(* Logix 5000 project; controller UOWHF Emulate 5570 rev 30.12; software revision 30.00; part 6 of 13 *)
(* tags used below, declared in another part *)
   UOWHF_Add_c : DINT;
   UOWHF_Msg : DINT[16];
   UOWHF_OutputMaxInd : DINT;
   UOWHF_Result : DINT[16];
(* MainProgram, continued *)

   		UOWHF_Result[5].31:=0;
   		UOWHF_Result[6]:=UOWHF_Result[6] + 895405157+UOWHF_Add_c;
   		UOWHF_Add_c.6:=UOWHF_Result[6].31;
   		UOWHF_Result[6].31:=0;
   	End_If;
   	If UOWHF_Msg[9].[21] Then
   		UOWHF_Result[0]:=UOWHF_Result[0] + 660161237+UOWHF_Add_c;
   		UOWHF_Add_c.0:=UOWHF_Result[0].31;
   		UOWHF_Result[0].31:=0;
   		UOWHF_Result[1]:=UOWHF_Result[1] + 1315089035+UOWHF_Add_c;
   		UOWHF_Add_c.1:=UOWHF_Result[1].31;
   		UOWHF_Result[1].31:=0;
   		UOWHF_Result[2]:=UOWHF_Result[2] + 1287512548+UOWHF_Add_c;
   		UOWHF_Add_c.2:=UOWHF_Result[2].31;
   		UOWHF_Result[2].31:=0;
   		UOWHF_Result[3]:=UOWHF_Result[3] + 1179731775+UOWHF_Add_c;
   		UOWHF_Add_c.3:=UOWHF_Result[3].31;
   		UOWHF_Result[3].31:=0;
   		UOWHF_Result[4]:=UOWHF_Result[4] + 1598255528+UOWHF_Add_c;
   		UOWHF_Add_c.4:=UOWHF_Result[4].31;
   		UOWHF_Result[4].31:=0;
   		UOWHF_Result[5]:=UOWHF_Result[5] + 1383999784+UOWHF_Add_c;
   		UOWHF_Add_c.5:=UOWHF_Result[5].31;
   		UOWHF_Result[5].31:=0;
   		UOWHF_Result[6]:=UOWHF_Result[6] + 83372341+UOWHF_Add_c;
   		UOWHF_Add_c.6:=UOWHF_Result[6].31;
   		UOWHF_Result[6].31:=0;
   	End_If;
   	If UOWHF_Msg[9].[22] Then
   		UOWHF_Result[0]:=UOWHF_Result[0] + 1715876547+UOWHF_Add_c;
   		UOWHF_Add_c.0:=UOWHF_Result[0].31;
   		UOWHF_Result[0].31:=0;
   		UOWHF_Result[1]:=UOWHF_Result[1] + 985647794+UOWHF_Add_c;
   		UOWHF_Add_c.1:=UOWHF_Result[1].31;
   		UOWHF_Result[1].31:=0;
   		UOWHF_Result[2]:=UOWHF_Result[2] + 1915071159+UOWHF_Add_c;
   		UOWHF_Add_c.2:=UOWHF_Result[2].31;
   		UOWHF_Result[2].31:=0;
   		UOWHF_Result[3]:=UOWHF_Result[3] + 1355115977+UOWHF_Add_c;
   		UOWHF_Add_c.3:=UOWHF_Result[3].31;
   		UOWHF_Result[3].31:=0;
   		UOWHF_Result[4]:=UOWHF_Result[4] + 296913181+UOWHF_Add_c;
   		UOWHF_Add_c.4:=UOWHF_Result[4].31;
   		UOWHF_Result[4].31:=0;
   		UOWHF_Result[5]:=UOWHF_Result[5] + 1237257487+UOWHF_Add_c;
   		UOWHF_Add_c.5:=UOWHF_Result[5].31;
   		UOWHF_Result[5].31:=0;
   		UOWHF_Result[6]:=UOWHF_Result[6] + 1778504117+UOWHF_Add_c;
   		UOWHF_Add_c.6:=UOWHF_Result[6].31;
   		UOWHF_Result[6].31:=0;
   	End_If;
   	If UOWHF_Msg[9].[23] Then
   		UOWHF_Result[0]:=UOWHF_Result[0] + 164662309+UOWHF_Add_c;
   		UOWHF_Add_c.0:=UOWHF_Result[0].31;
   		UOWHF_Result[0].31:=0;
   		UOWHF_Result[1]:=UOWHF_Result[1] + 1325365703+UOWHF_Add_c;
   		UOWHF_Add_c.1:=UOWHF_Result[1].31;
   		UOWHF_Result[1].31:=0;
   		UOWHF_Result[2]:=UOWHF_Result[2] + 1493283531+UOWHF_Add_c;
   		UOWHF_Add_c.2:=UOWHF_Result[2].31;
   		UOWHF_Result[2].31:=0;
   		UOWHF_Result[3]:=UOWHF_Result[3] + 2135510542+UOWHF_Add_c;
   		UOWHF_Add_c.3:=UOWHF_Result[3].31;
   		UOWHF_Result[3].31:=0;
   		UOWHF_Result[4]:=UOWHF_Result[4] + 1163293199+UOWHF_Add_c;
   		UOWHF_Add_c.4:=UOWHF_Result[4].31;
   		UOWHF_Result[4].31:=0;
   		UOWHF_Result[5]:=UOWHF_Result[5] + 92683402+UOWHF_Add_c;
   		UOWHF_Add_c.5:=UOWHF_Result[5].31;
   		UOWHF_Result[5].31:=0;
   		UOWHF_Result[6]:=UOWHF_Result[6] + 1965230931+UOWHF_Add_c;
   		UOWHF_Add_c.6:=UOWHF_Result[6].31;
   		UOWHF_Result[6].31:=0;
   	End_If;
   	If UOWHF_Msg[9].[24] Then
   		UOWHF_Result[0]:=UOWHF_Result[0] + 1349986349+UOWHF_Add_c;
   		UOWHF_Add_c.0:=UOWHF_Result[0].31;
   		UOWHF_Result[0].31:=0;
   		UOWHF_Result[1]:=UOWHF_Result[1] + 1428111799+UOWHF_Add_c;
   		UOWHF_Add_c.1:=UOWHF_Result[1].31;
   		UOWHF_Result[1].31:=0;
   		UOWHF_Result[2]:=UOWHF_Result[2] + 168351548+UOWHF_Add_c;
   		UOWHF_Add_c.2:=UOWHF_Result[2].31;
   		UOWHF_Result[2].31:=0;
   		UOWHF_Result[3]:=UOWHF_Result[3] + 1291854191+UOWHF_Add_c;
   		UOWHF_Add_c.3:=UOWHF_Result[3].31;
   		UOWHF_Result[3].31:=0;
   		UOWHF_Result[4]:=UOWHF_Result[4] + 1544153517+UOWHF_Add_c;
   		UOWHF_Add_c.4:=UOWHF_Result[4].31;
   		UOWHF_Result[4].31:=0;
   		UOWHF_Result[5]:=UOWHF_Result[5] + 1624211329+UOWHF_Add_c;
   		UOWHF_Add_c.5:=UOWHF_Result[5].31;
   		UOWHF_Result[5].31:=0;
   		UOWHF_Result[6]:=UOWHF_Result[6] + 1832912649+UOWHF_Add_c;
   		UOWHF_Add_c.6:=UOWHF_Result[6].31;
   		UOWHF_Result[6].31:=0;
   	End_If;
   	If UOWHF_Msg[9].[25] Then
   		UOWHF_Result[0]:=UOWHF_Result[0] + 1267672492+UOWHF_Add_c;
   		UOWHF_Add_c.0:=UOWHF_Result[0].31;
   		UOWHF_Result[0].31:=0;
   		UOWHF_Result[1]:=UOWHF_Result[1] + 884086529+UOWHF_Add_c;
   		UOWHF_Add_c.1:=UOWHF_Result[1].31;
   		UOWHF_Result[1].31:=0;
   		UOWHF_Result[2]:=UOWHF_Result[2] + 1230680266+UOWHF_Add_c;
   		UOWHF_Add_c.2:=UOWHF_Result[2].31;
   		UOWHF_Result[2].31:=0;
   		UOWHF_Result[3]:=UOWHF_Result[3] + 485350037+UOWHF_Add_c;
   		UOWHF_Add_c.3:=UOWHF_Result[3].31;
   		UOWHF_Result[3].31:=0;
   		UOWHF_Result[4]:=UOWHF_Result[4] + 1714826949+UOWHF_Add_c;
   		UOWHF_Add_c.4:=UOWHF_Result[4].31;
   		UOWHF_Result[4].31:=0;
   		UOWHF_Result[5]:=UOWHF_Result[5] + 1853366658+UOWHF_Add_c;
   		UOWHF_Add_c.5:=UOWHF_Result[5].31;
   		UOWHF_Result[5].31:=0;
   		UOWHF_Result[6]:=UOWHF_Result[6] + 1466072212+UOWHF_Add_c;
   		UOWHF_Add_c.6:=UOWHF_Result[6].31;
   		UOWHF_Result[6].31:=0;
   	End_If;
   	If UOWHF_Msg[9].[26] Then
   		UOWHF_Result[0]:=UOWHF_Result[0] + 755970944+UOWHF_Add_c;
   		UOWHF_Add_c.0:=UOWHF_Result[0].31;
   		UOWHF_Result[0].31:=0;
   		UOWHF_Result[1]:=UOWHF_Result[1] + 2084777862+UOWHF_Add_c;
   		UOWHF_Add_c.1:=UOWHF_Result[1].31;
   		UOWHF_Result[1].31:=0;
   		UOWHF_Result[2]:=UOWHF_Result[2] + 328525721+UOWHF_Add_c;
   		UOWHF_Add_c.2:=UOWHF_Result[2].31;
   		UOWHF_Result[2].31:=0;
   		UOWHF_Result[3]:=UOWHF_Result[3] + 1005208267+UOWHF_Add_c;
   		UOWHF_Add_c.3:=UOWHF_Result[3].31;
   		UOWHF_Result[3].31:=0;
   		UOWHF_Result[4]:=UOWHF_Result[4] + 1410939800+UOWHF_Add_c;
   		UOWHF_Add_c.4:=UOWHF_Result[4].31;
   		UOWHF_Result[4].31:=0;
   		UOWHF_Result[5]:=UOWHF_Result[5] + 813260174+UOWHF_Add_c;
   		UOWHF_Add_c.5:=UOWHF_Result[5].31;
   		UOWHF_Result[5].31:=0;
   		UOWHF_Result[6]:=UOWHF_Result[6] + 547964095+UOWHF_Add_c;
   		UOWHF_Add_c.6:=UOWHF_Result[6].31;
   		UOWHF_Result[6].31:=0;
   	End_If;
   	If UOWHF_Msg[9].[27] Then
   		UOWHF_Result[0]:=UOWHF_Result[0] + 997423673+UOWHF_Add_c;
   		UOWHF_Add_c.0:=UOWHF_Result[0].31;
   		UOWHF_Result[0].31:=0;
   		UOWHF_Result[1]:=UOWHF_Result[1] + 1791173720+UOWHF_Add_c;
   		UOWHF_Add_c.1:=UOWHF_Result[1].31;
   		UOWHF_Result[1].31:=0;
   		UOWHF_Result[2]:=UOWHF_Result[2] + 466501049+UOWHF_Add_c;
   		UOWHF_Add_c.2:=UOWHF_Result[2].31;
   		UOWHF_Result[2].31:=0;
   		UOWHF_Result[3]:=UOWHF_Result[3] + 1763922528+UOWHF_Add_c;
   		UOWHF_Add_c.3:=UOWHF_Result[3].31;
   		UOWHF_Result[3].31:=0;
   		UOWHF_Result[4]:=UOWHF_Result[4] + 1977911472+UOWHF_Add_c;
   		UOWHF_Add_c.4:=UOWHF_Result[4].31;
   		UOWHF_Result[4].31:=0;
   		UOWHF_Result[5]:=UOWHF_Result[5] + 1301488429+UOWHF_Add_c;
   		UOWHF_Add_c.5:=UOWHF_Result[5].31;
   		UOWHF_Result[5].31:=0;
   		UOWHF_Result[6]:=UOWHF_Result[6] + 1196244772+UOWHF_Add_c;
   		UOWHF_Add_c.6:=UOWHF_Result[6].31;
   		UOWHF_Result[6].31:=0;
   	End_If;
   	If UOWHF_Msg[9].[28] Then
   		UOWHF_Result[0]:=UOWHF_Result[0] + 1877124502+UOWHF_Add_c;
   		UOWHF_Add_c.0:=UOWHF_Result[0].31;
   		UOWHF_Result[0].31:=0;
   		UOWHF_Result[1]:=UOWHF_Result[1] + 1015259037+UOWHF_Add_c;
   		UOWHF_Add_c.1:=UOWHF_Result[1].31;
   		UOWHF_Result[1].31:=0;
   		UOWHF_Result[2]:=UOWHF_Result[2] + 1954515831+UOWHF_Add_c;
   		UOWHF_Add_c.2:=UOWHF_Result[2].31;
   		UOWHF_Result[2].31:=0;
   		UOWHF_Result[3]:=UOWHF_Result[3] + 1806236750+UOWHF_Add_c;
   		UOWHF_Add_c.3:=UOWHF_Result[3].31;
   		UOWHF_Result[3].31:=0;
   		UOWHF_Result[4]:=UOWHF_Result[4] + 458134772+UOWHF_Add_c;
   		UOWHF_Add_c.4:=UOWHF_Result[4].31;
   		UOWHF_Result[4].31:=0;
   		UOWHF_Result[5]:=UOWHF_Result[5] + 419069533+UOWHF_Add_c;
   		UOWHF_Add_c.5:=UOWHF_Result[5].31;
   		UOWHF_Result[5].31:=0;
   		UOWHF_Result[6]:=UOWHF_Result[6] + 790941477+UOWHF_Add_c;
   		UOWHF_Add_c.6:=UOWHF_Result[6].31;
   		UOWHF_Result[6].31:=0;
   	End_If;
   	If UOWHF_Msg[9].[29] Then
   		UOWHF_Result[0]:=UOWHF_Result[0] + 1874899523+UOWHF_Add_c;
   		UOWHF_Add_c.0:=UOWHF_Result[0].31;
   		UOWHF_Result[0].31:=0;
   		UOWHF_Result[1]:=UOWHF_Result[1] + 1348598912+UOWHF_Add_c;
   		UOWHF_Add_c.1:=UOWHF_Result[1].31;
   		UOWHF_Result[1].31:=0;
   		UOWHF_Result[2]:=UOWHF_Result[2] + 2101684580+UOWHF_Add_c;
   		UOWHF_Add_c.2:=UOWHF_Result[2].31;
   		UOWHF_Result[2].31:=0;
   		UOWHF_Result[3]:=UOWHF_Result[3] + 1884890663+UOWHF_Add_c;
   		UOWHF_Add_c.3:=UOWHF_Result[3].31;
   		UOWHF_Result[3].31:=0;
   		UOWHF_Result[4]:=UOWHF_Result[4] + 1188937122+UOWHF_Add_c;
   		UOWHF_Add_c.4:=UOWHF_Result[4].31;
   		UOWHF_Result[4].31:=0;
   		UOWHF_Result[5]:=UOWHF_Result[5] + 2029021445+UOWHF_Add_c;
   		UOWHF_Add_c.5:=UOWHF_Result[5].31;
   		UOWHF_Result[5].31:=0;
   		UOWHF_Result[6]:=UOWHF_Result[6] + 1538909396+UOWHF_Add_c;
   		UOWHF_Add_c.6:=UOWHF_Result[6].31;
   		UOWHF_Result[6].31:=0;
   	End_If;
   	If UOWHF_Msg[9].[30] Then
   		UOWHF_Result[0]:=UOWHF_Result[0] + 235965658+UOWHF_Add_c;
   		UOWHF_Add_c.0:=UOWHF_Result[0].31;
   		UOWHF_Result[0].31:=0;
   		UOWHF_Result[1]:=UOWHF_Result[1] + 1317732388+UOWHF_Add_c;
   		UOWHF_Add_c.1:=UOWHF_Result[1].31;
   		UOWHF_Result[1].31:=0;
   		UOWHF_Result[2]:=UOWHF_Result[2] + 1030092944+UOWHF_Add_c;
   		UOWHF_Add_c.2:=UOWHF_Result[2].31;
   		UOWHF_Result[2].31:=0;
   		UOWHF_Result[3]:=UOWHF_Result[3] + 1908438518+UOWHF_Add_c;
   		UOWHF_Add_c.3:=UOWHF_Result[3].31;
   		UOWHF_Result[3].31:=0;
   		UOWHF_Result[4]:=UOWHF_Result[4] + 919181552+UOWHF_Add_c;
   		UOWHF_Add_c.4:=UOWHF_Result[4].31;
   		UOWHF_Result[4].31:=0;
   		UOWHF_Result[5]:=UOWHF_Result[5] + 239215457+UOWHF_Add_c;
   		UOWHF_Add_c.5:=UOWHF_Result[5].31;
   		UOWHF_Result[5].31:=0;
   		UOWHF_Result[6]:=UOWHF_Result[6] + 1472128231+UOWHF_Add_c;
   		UOWHF_Add_c.6:=UOWHF_Result[6].31;
   		UOWHF_Result[6].31:=0;
   	End_If;
   	If UOWHF_Msg[9].[31] Then
   		UOWHF_Result[0]:=UOWHF_Result[0] + 1398442323+UOWHF_Add_c;
   		UOWHF_Add_c.0:=UOWHF_Result[0].31;
   		UOWHF_Result[0].31:=0;
   		UOWHF_Result[1]:=UOWHF_Result[1] + 964623714+UOWHF_Add_c;
   		UOWHF_Add_c.1:=UOWHF_Result[1].31;
   		UOWHF_Result[1].31:=0;
   		UOWHF_Result[2]:=UOWHF_Result[2] + 256294152+UOWHF_Add_c;
   		UOWHF_Add_c.2:=UOWHF_Result[2].31;
   		UOWHF_Result[2].31:=0;
   		UOWHF_Result[3]:=UOWHF_Result[3] + 1907160525+UOWHF_Add_c;
   		UOWHF_Add_c.3:=UOWHF_Result[3].31;
   		UOWHF_Result[3].31:=0;
   		UOWHF_Result[4]:=UOWHF_Result[4] + 846515090+UOWHF_Add_c;
   		UOWHF_Add_c.4:=UOWHF_Result[4].31;
   		UOWHF_Result[4].31:=0;
   		UOWHF_Result[5]:=UOWHF_Result[5] + 958207881+UOWHF_Add_c;
   		UOWHF_Add_c.5:=UOWHF_Result[5].31;
   		UOWHF_Result[5].31:=0;
   		UOWHF_Result[6]:=UOWHF_Result[6] + 1865822718+UOWHF_Add_c;
   		UOWHF_Add_c.6:=UOWHF_Result[6].31;
   		UOWHF_Result[6].31:=0;
   	End_If;
   	If UOWHF_Msg[10].[0] Then
   		UOWHF_Result[0]:=UOWHF_Result[0] + 1543145221+UOWHF_Add_c;
   		UOWHF_Add_c.0:=UOWHF_Result[0].31;
   		UOWHF_Result[0].31:=0;
   		UOWHF_Result[1]:=UOWHF_Result[1] + 1596571495+UOWHF_Add_c;
   		UOWHF_Add_c.1:=UOWHF_Result[1].31;
   		UOWHF_Result[1].31:=0;
   		UOWHF_Result[2]:=UOWHF_Result[2] + 1603169829+UOWHF_Add_c;
   		UOWHF_Add_c.2:=UOWHF_Result[2].31;
   		UOWHF_Result[2].31:=0;
   		UOWHF_Result[3]:=UOWHF_Result[3] + 2046965193+UOWHF_Add_c;
   		UOWHF_Add_c.3:=UOWHF_Result[3].31;
   		UOWHF_Result[3].31:=0;
   		UOWHF_Result[4]:=UOWHF_Result[4] + 1757211017+UOWHF_Add_c;
   		UOWHF_Add_c.4:=UOWHF_Result[4].31;
   		UOWHF_Result[4].31:=0;
   		UOWHF_Result[5]:=UOWHF_Result[5] + 130098380+UOWHF_Add_c;
   		UOWHF_Add_c.5:=UOWHF_Result[5].31;
   		UOWHF_Result[5].31:=0;
   		UOWHF_Result[6]:=UOWHF_Result[6] + 1310384925+UOWHF_Add_c;
   		UOWHF_Add_c.6:=UOWHF_Result[6].31;
   		UOWHF_Result[6].31:=0;
   	End_If;
   	If UOWHF_Msg[10].[1] Then
   		UOWHF_Result[0]:=UOWHF_Result[0] + 126953638+UOWHF_Add_c;
   		UOWHF_Add_c.0:=UOWHF_Result[0].31;
   		UOWHF_Result[0].31:=0;
   		UOWHF_Result[1]:=UOWHF_Result[1] + 1013212484+UOWHF_Add_c;
   		UOWHF_Add_c.1:=UOWHF_Result[1].31;
   		UOWHF_Result[1].31:=0;
   		UOWHF_Result[2]:=UOWHF_Result[2] + 815619305+UOWHF_Add_c;
   		UOWHF_Add_c.2:=UOWHF_Result[2].31;
   		UOWHF_Result[2].31:=0;
   		UOWHF_Result[3]:=UOWHF_Result[3] + 677856911+UOWHF_Add_c;
   		UOWHF_Add_c.3:=UOWHF_Result[3].31;
   		UOWHF_Result[3].31:=0;
   		UOWHF_Result[4]:=UOWHF_Result[4] + 1261957295+UOWHF_Add_c;
   		UOWHF_Add_c.4:=UOWHF_Result[4].31;
   		UOWHF_Result[4].31:=0;
   		UOWHF_Result[5]:=UOWHF_Result[5] + 1834778391+UOWHF_Add_c;
   		UOWHF_Add_c.5:=UOWHF_Result[5].31;
   		UOWHF_Result[5].31:=0;
   		UOWHF_Result[6]:=UOWHF_Result[6] + 167047653+UOWHF_Add_c;
   		UOWHF_Add_c.6:=UOWHF_Result[6].31;
   		UOWHF_Result[6].31:=0;
   	End_If;
   	If UOWHF_Msg[10].[2] Then
   		UOWHF_Result[0]:=UOWHF_Result[0] + 1265210804+UOWHF_Add_c;
   		UOWHF_Add_c.0:=UOWHF_Result[0].31;
   		UOWHF_Result[0].31:=0;
   		UOWHF_Result[1]:=UOWHF_Result[1] + 940847770+UOWHF_Add_c;
   		UOWHF_Add_c.1:=UOWHF_Result[1].31;
   		UOWHF_Result[1].31:=0;
   		UOWHF_Result[2]:=UOWHF_Result[2] + 969325259+UOWHF_Add_c;
   		UOWHF_Add_c.2:=UOWHF_Result[2].31;
   		UOWHF_Result[2].31:=0;
   		UOWHF_Result[3]:=UOWHF_Result[3] + 367906621+UOWHF_Add_c;
   		UOWHF_Add_c.3:=UOWHF_Result[3].31;
   		UOWHF_Result[3].31:=0;
   		UOWHF_Result[4]:=UOWHF_Result[4] + 1871994288+UOWHF_Add_c;
   		UOWHF_Add_c.4:=UOWHF_Result[4].31;
   		UOWHF_Result[4].31:=0;
   		UOWHF_Result[5]:=UOWHF_Result[5] + 638431925+UOWHF_Add_c;
   		UOWHF_Add_c.5:=UOWHF_Result[5].31;
   		UOWHF_Result[5].31:=0;
   		UOWHF_Result[6]:=UOWHF_Result[6] + 994996741+UOWHF_Add_c;
   		UOWHF_Add_c.6:=UOWHF_Result[6].31;
   		UOWHF_Result[6].31:=0;
   	End_If;
   	If UOWHF_Msg[10].[3] Then
   		UOWHF_Result[0]:=UOWHF_Result[0] + 1816124282+UOWHF_Add_c;
   		UOWHF_Add_c.0:=UOWHF_Result[0].31;
   		UOWHF_Result[0].31:=0;
   		UOWHF_Result[1]:=UOWHF_Result[1] + 1763814085+UOWHF_Add_c;
   		UOWHF_Add_c.1:=UOWHF_Result[1].31;
   		UOWHF_Result[1].31:=0;
   		UOWHF_Result[2]:=UOWHF_Result[2] + 2035926671+UOWHF_Add_c;
   		UOWHF_Add_c.2:=UOWHF_Result[2].31;
   		UOWHF_Result[2].31:=0;
   		UOWHF_Result[3]:=UOWHF_Result[3] + 591419378+UOWHF_Add_c;
   		UOWHF_Add_c.3:=UOWHF_Result[3].31;
   		UOWHF_Result[3].31:=0;
   		UOWHF_Result[4]:=UOWHF_Result[4] + 1709863160+UOWHF_Add_c;
   		UOWHF_Add_c.4:=UOWHF_Result[4].31;
   		UOWHF_Result[4].31:=0;
   		UOWHF_Result[5]:=UOWHF_Result[5] + 2133800064+UOWHF_Add_c;
   		UOWHF_Add_c.5:=UOWHF_Result[5].31;
   		UOWHF_Result[5].31:=0;
   		UOWHF_Result[6]:=UOWHF_Result[6] + 1339032441+UOWHF_Add_c;
   		UOWHF_Add_c.6:=UOWHF_Result[6].31;
   		UOWHF_Result[6].31:=0;
   	End_If;
   	If UOWHF_Msg[10].[4] Then
   		UOWHF_Result[0]:=UOWHF_Result[0] + 854930131+UOWHF_Add_c;
   		UOWHF_Add_c.0:=UOWHF_Result[0].31;
   		UOWHF_Result[0].31:=0;
   		UOWHF_Result[1]:=UOWHF_Result[1] + 1372200423+UOWHF_Add_c;
   		UOWHF_Add_c.1:=UOWHF_Result[1].31;
   		UOWHF_Result[1].31:=0;
   		UOWHF_Result[2]:=UOWHF_Result[2] + 2131196727+UOWHF_Add_c;
   		UOWHF_Add_c.2:=UOWHF_Result[2].31;
   		UOWHF_Result[2].31:=0;
   		UOWHF_Result[3]:=UOWHF_Result[3] + 853135064+UOWHF_Add_c;
   		UOWHF_Add_c.3:=UOWHF_Result[3].31;
   		UOWHF_Result[3].31:=0;
   		UOWHF_Result[4]:=UOWHF_Result[4] + 1495256040+UOWHF_Add_c;
   		UOWHF_Add_c.4:=UOWHF_Result[4].31;
   		UOWHF_Result[4].31:=0;
   		UOWHF_Result[5]:=UOWHF_Result[5] + 222151544+UOWHF_Add_c;
   		UOWHF_Add_c.5:=UOWHF_Result[5].31;
   		UOWHF_Result[5].31:=0;
   		UOWHF_Result[6]:=UOWHF_Result[6] + 754259260+UOWHF_Add_c;
   		UOWHF_Add_c.6:=UOWHF_Result[6].31;
   		UOWHF_Result[6].31:=0;
   	End_If;
   	If UOWHF_Msg[10].[5] Then
   		UOWHF_Result[0]:=UOWHF_Result[0] + 1563421875+UOWHF_Add_c;
   		UOWHF_Add_c.0:=UOWHF_Result[0].31;
   		UOWHF_Result[0].31:=0;
   		UOWHF_Result[1]:=UOWHF_Result[1] + 242182278+UOWHF_Add_c;
   		UOWHF_Add_c.1:=UOWHF_Result[1].31;
   		UOWHF_Result[1].31:=0;
   		UOWHF_Result[2]:=UOWHF_Result[2] + 436664119+UOWHF_Add_c;
   		UOWHF_Add_c.2:=UOWHF_Result[2].31;
   		UOWHF_Result[2].31:=0;
   		UOWHF_Result[3]:=UOWHF_Result[3] + 1075520283+UOWHF_Add_c;
   		UOWHF_Add_c.3:=UOWHF_Result[3].31;
   		UOWHF_Result[3].31:=0;
   		UOWHF_Result[4]:=UOWHF_Result[4] + 448912110+UOWHF_Add_c;
   		UOWHF_Add_c.4:=UOWHF_Result[4].31;
   		UOWHF_Result[4].31:=0;
   		UOWHF_Result[5]:=UOWHF_Result[5] + 1908828426+UOWHF_Add_c;
   		UOWHF_Add_c.5:=UOWHF_Result[5].31;
   		UOWHF_Result[5].31:=0;
   		UOWHF_Result[6]:=UOWHF_Result[6] + 1950510765+UOWHF_Add_c;
   		UOWHF_Add_c.6:=UOWHF_Result[6].31;
   		UOWHF_Result[6].31:=0;
   	End_If;
   	If UOWHF_Msg[10].[6] Then
   		UOWHF_Result[0]:=UOWHF_Result[0] + 624941020+UOWHF_Add_c;
   		UOWHF_Add_c.0:=UOWHF_Result[0].31;
   		UOWHF_Result[0].31:=0;
   		UOWHF_Result[1]:=UOWHF_Result[1] + 1171201426+UOWHF_Add_c;
   		UOWHF_Add_c.1:=UOWHF_Result[1].31;
   		UOWHF_Result[1].31:=0;
   		UOWHF_Result[2]:=UOWHF_Result[2] + 537642592+UOWHF_Add_c;
   		UOWHF_Add_c.2:=UOWHF_Result[2].31;
   		UOWHF_Result[2].31:=0;
   		UOWHF_Result[3]:=UOWHF_Result[3] + 420524488+UOWHF_Add_c;
   		UOWHF_Add_c.3:=UOWHF_Result[3].31;
   		UOWHF_Result[3].31:=0;
   		UOWHF_Result[4]:=UOWHF_Result[4] + 477664528+UOWHF_Add_c;
   		UOWHF_Add_c.4:=UOWHF_Result[4].31;
   		UOWHF_Result[4].31:=0;
   		UOWHF_Result[5]:=UOWHF_Result[5] + 362505463+UOWHF_Add_c;
   		UOWHF_Add_c.5:=UOWHF_Result[5].31;
   		UOWHF_Result[5].31:=0;
   		UOWHF_Result[6]:=UOWHF_Result[6] + 1995831580+UOWHF_Add_c;
   		UOWHF_Add_c.6:=UOWHF_Result[6].31;
   		UOWHF_Result[6].31:=0;
   	End_If;
   	If UOWHF_Msg[10].[7] Then
   		UOWHF_Result[0]:=UOWHF_Result[0] + 1657679202+UOWHF_Add_c;
   		UOWHF_Add_c.0:=UOWHF_Result[0].31;
   		UOWHF_Result[0].31:=0;
   		UOWHF_Result[1]:=UOWHF_Result[1] + 1342754235+UOWHF_Add_c;
   		UOWHF_Add_c.1:=UOWHF_Result[1].31;
   		UOWHF_Result[1].31:=0;
   		UOWHF_Result[2]:=UOWHF_Result[2] + 1471900463+UOWHF_Add_c;
   		UOWHF_Add_c.2:=UOWHF_Result[2].31;
   		UOWHF_Result[2].31:=0;
   		UOWHF_Result[3]:=UOWHF_Result[3] + 1684834987+UOWHF_Add_c;
   		UOWHF_Add_c.3:=UOWHF_Result[3].31;
   		UOWHF_Result[3].31:=0;
   		UOWHF_Result[4]:=UOWHF_Result[4] + 1214737626+UOWHF_Add_c;
   		UOWHF_Add_c.4:=UOWHF_Result[4].31;
   		UOWHF_Result[4].31:=0;
   		UOWHF_Result[5]:=UOWHF_Result[5] + 1907134264+UOWHF_Add_c;
   		UOWHF_Add_c.5:=UOWHF_Result[5].31;
   		UOWHF_Result[5].31:=0;
   		UOWHF_Result[6]:=UOWHF_Result[6] + 1587406036+UOWHF_Add_c;
   		UOWHF_Add_c.6:=UOWHF_Result[6].31;
   		UOWHF_Result[6].31:=0;
   	End_If;
   	If UOWHF_Msg[10].[8] Then
   		UOWHF_Result[0]:=UOWHF_Result[0] + 526080272+UOWHF_Add_c;
   		UOWHF_Add_c.0:=UOWHF_Result[0].31;
   		UOWHF_Result[0].31:=0;
   		UOWHF_Result[1]:=UOWHF_Result[1] + 362791028+UOWHF_Add_c;
   		UOWHF_Add_c.1:=UOWHF_Result[1].31;
   		UOWHF_Result[1].31:=0;
   		UOWHF_Result[2]:=UOWHF_Result[2] + 1719461918+UOWHF_Add_c;
   		UOWHF_Add_c.2:=UOWHF_Result[2].31;
   		UOWHF_Result[2].31:=0;
   		UOWHF_Result[3]:=UOWHF_Result[3] + 427154490+UOWHF_Add_c;
   		UOWHF_Add_c.3:=UOWHF_Result[3].31;
   		UOWHF_Result[3].31:=0;
   		UOWHF_Result[4]:=UOWHF_Result[4] + 798716505+UOWHF_Add_c;
   		UOWHF_Add_c.4:=UOWHF_Result[4].31;
   		UOWHF_Result[4].31:=0;
   		UOWHF_Result[5]:=UOWHF_Result[5] + 690658399+UOWHF_Add_c;
   		UOWHF_Add_c.5:=UOWHF_Result[5].31;
   		UOWHF_Result[5].31:=0;
   		UOWHF_Result[6]:=UOWHF_Result[6] + 399269664+UOWHF_Add_c;
   		UOWHF_Add_c.6:=UOWHF_Result[6].31;
   		UOWHF_Result[6].31:=0;
   	End_If;
   	If UOWHF_Msg[10].[9] Then
   		UOWHF_Result[0]:=UOWHF_Result[0] + 2107724001+UOWHF_Add_c;
   		UOWHF_Add_c.0:=UOWHF_Result[0].31;
   		UOWHF_Result[0].31:=0;
   		UOWHF_Result[1]:=UOWHF_Result[1] + 1057490839+UOWHF_Add_c;
   		UOWHF_Add_c.1:=UOWHF_Result[1].31;
   		UOWHF_Result[1].31:=0;
   		UOWHF_Result[2]:=UOWHF_Result[2] + 879111903+UOWHF_Add_c;
   		UOWHF_Add_c.2:=UOWHF_Result[2].31;
   		UOWHF_Result[2].31:=0;
   		UOWHF_Result[3]:=UOWHF_Result[3] + 1230271781+UOWHF_Add_c;
   		UOWHF_Add_c.3:=UOWHF_Result[3].31;
   		UOWHF_Result[3].31:=0;
   		UOWHF_Result[4]:=UOWHF_Result[4] + 238135446+UOWHF_Add_c;
   		UOWHF_Add_c.4:=UOWHF_Result[4].31;
   		UOWHF_Result[4].31:=0;
   		UOWHF_Result[5]:=UOWHF_Result[5] + 1989397853+UOWHF_Add_c;
   		UOWHF_Add_c.5:=UOWHF_Result[5].31;
   		UOWHF_Result[5].31:=0;
   		UOWHF_Result[6]:=UOWHF_Result[6] + 1849353930+UOWHF_Add_c;
   		UOWHF_Add_c.6:=UOWHF_Result[6].31;
   		UOWHF_Result[6].31:=0;
   	End_If;
   	If UOWHF_Msg[10].[10] Then
   		UOWHF_Result[0]:=UOWHF_Result[0] + 918739460+UOWHF_Add_c;
   		UOWHF_Add_c.0:=UOWHF_Result[0].31;
   		UOWHF_Result[0].31:=0;
   		UOWHF_Result[1]:=UOWHF_Result[1] + 1059272652+UOWHF_Add_c;
   		UOWHF_Add_c.1:=UOWHF_Result[1].31;
   		UOWHF_Result[1].31:=0;
   		UOWHF_Result[2]:=UOWHF_Result[2] + 1378794548+UOWHF_Add_c;
   		UOWHF_Add_c.2:=UOWHF_Result[2].31;
   		UOWHF_Result[2].31:=0;
   		UOWHF_Result[3]:=UOWHF_Result[3] + 2021810889+UOWHF_Add_c;
   		UOWHF_Add_c.3:=UOWHF_Result[3].31;
   		UOWHF_Result[3].31:=0;
   		UOWHF_Result[4]:=UOWHF_Result[4] + 2124083835+UOWHF_Add_c;
   		UOWHF_Add_c.4:=UOWHF_Result[4].31;
   		UOWHF_Result[4].31:=0;
   		UOWHF_Result[5]:=UOWHF_Result[5] + 1555199521+UOWHF_Add_c;
   		UOWHF_Add_c.5:=UOWHF_Result[5].31;
   		UOWHF_Result[5].31:=0;
   		UOWHF_Result[6]:=UOWHF_Result[6] + 1959982309+UOWHF_Add_c;
   		UOWHF_Add_c.6:=UOWHF_Result[6].31;
   		UOWHF_Result[6].31:=0;
   	End_If;
   	If UOWHF_Msg[10].[11] Then
   		UOWHF_Result[0]:=UOWHF_Result[0] + 409848939+UOWHF_Add_c;
   		UOWHF_Add_c.0:=UOWHF_Result[0].31;
   		UOWHF_Result[0].31:=0;
   		UOWHF_Result[1]:=UOWHF_Result[1] + 2000970897+UOWHF_Add_c;
   		UOWHF_Add_c.1:=UOWHF_Result[1].31;
   		UOWHF_Result[1].31:=0;
   		UOWHF_Result[2]:=UOWHF_Result[2] + 577580939+UOWHF_Add_c;
   		UOWHF_Add_c.2:=UOWHF_Result[2].31;
   		UOWHF_Result[2].31:=0;
   		UOWHF_Result[3]:=UOWHF_Result[3] + 1672799932+UOWHF_Add_c;
   		UOWHF_Add_c.3:=UOWHF_Result[3].31;
   		UOWHF_Result[3].31:=0;
   		UOWHF_Result[4]:=UOWHF_Result[4] + 2115458545+UOWHF_Add_c;
   		UOWHF_Add_c.4:=UOWHF_Result[4].31;
   		UOWHF_Result[4].31:=0;
   		UOWHF_Result[5]:=UOWHF_Result[5] + 1030388630+UOWHF_Add_c;
   		UOWHF_Add_c.5:=UOWHF_Result[5].31;
   		UOWHF_Result[5].31:=0;
   		UOWHF_Result[6]:=UOWHF_Result[6] + 1934563828+UOWHF_Add_c;
   		UOWHF_Add_c.6:=UOWHF_Result[6].31;
   		UOWHF_Result[6].31:=0;
   	End_If;
   	If UOWHF_Msg[10].[12] Then
   		UOWHF_Result[0]:=UOWHF_Result[0] + 376288360+UOWHF_Add_c;
   		UOWHF_Add_c.0:=UOWHF_Result[0].31;
   		UOWHF_Result[0].31:=0;
   		UOWHF_Result[1]:=UOWHF_Result[1] + 1208467327+UOWHF_Add_c;
   		UOWHF_Add_c.1:=UOWHF_Result[1].31;
   		UOWHF_Result[1].31:=0;
   		UOWHF_Result[2]:=UOWHF_Result[2] + 148525877+UOWHF_Add_c;
   		UOWHF_Add_c.2:=UOWHF_Result[2].31;
   		UOWHF_Result[2].31:=0;
   		UOWHF_Result[3]:=UOWHF_Result[3] + 896227724+UOWHF_Add_c;
   		UOWHF_Add_c.3:=UOWHF_Result[3].31;
   		UOWHF_Result[3].31:=0;
   		UOWHF_Result[4]:=UOWHF_Result[4] + 358257308+UOWHF_Add_c;
   		UOWHF_Add_c.4:=UOWHF_Result[4].31;
   		UOWHF_Result[4].31:=0;
   		UOWHF_Result[5]:=UOWHF_Result[5] + 126124772+UOWHF_Add_c;
   		UOWHF_Add_c.5:=UOWHF_Result[5].31;
   		UOWHF_Result[5].31:=0;
   		UOWHF_Result[6]:=UOWHF_Result[6] + 1944566+UOWHF_Add_c;
   		UOWHF_Add_c.6:=UOWHF_Result[6].31;
   		UOWHF_Result[6].31:=0;
   	End_If;
   	If UOWHF_Msg[10].[13] Then
   		UOWHF_Result[0]:=UOWHF_Result[0] + 1113461694+UOWHF_Add_c;
   		UOWHF_Add_c.0:=UOWHF_Result[0].31;
   		UOWHF_Result[0].31:=0;
   		UOWHF_Result[1]:=UOWHF_Result[1] + 37995443+UOWHF_Add_c;
   		UOWHF_Add_c.1:=UOWHF_Result[1].31;
   		UOWHF_Result[1].31:=0;
   		UOWHF_Result[2]:=UOWHF_Result[2] + 1197929973+UOWHF_Add_c;
   		UOWHF_Add_c.2:=UOWHF_Result[2].31;
   		UOWHF_Result[2].31:=0;
   		UOWHF_Result[3]:=UOWHF_Result[3] + 942197906+UOWHF_Add_c;
   		UOWHF_Add_c.3:=UOWHF_Result[3].31;
   		UOWHF_Result[3].31:=0;
   		UOWHF_Result[4]:=UOWHF_Result[4] + 894318581+UOWHF_Add_c;
   		UOWHF_Add_c.4:=UOWHF_Result[4].31;
   		UOWHF_Result[4].31:=0;
   		UOWHF_Result[5]:=UOWHF_Result[5] + 1370002959+UOWHF_Add_c;
   		UOWHF_Add_c.5:=UOWHF_Result[5].31;
   		UOWHF_Result[5].31:=0;
   		UOWHF_Result[6]:=UOWHF_Result[6] + 1796314076+UOWHF_Add_c;
   		UOWHF_Add_c.6:=UOWHF_Result[6].31;
   		UOWHF_Result[6].31:=0;
   	End_If;
   	If UOWHF_Msg[10].[14] Then
   		UOWHF_Result[0]:=UOWHF_Result[0] + 1569257492+UOWHF_Add_c;
   		UOWHF_Add_c.0:=UOWHF_Result[0].31;
   		UOWHF_Result[0].31:=0;
   		UOWHF_Result[1]:=UOWHF_Result[1] + 635645250+UOWHF_Add_c;
   		UOWHF_Add_c.1:=UOWHF_Result[1].31;
   		UOWHF_Result[1].31:=0;
   		UOWHF_Result[2]:=UOWHF_Result[2] + 2086282355+UOWHF_Add_c;
   		UOWHF_Add_c.2:=UOWHF_Result[2].31;
   		UOWHF_Result[2].31:=0;
   		UOWHF_Result[3]:=UOWHF_Result[3] + 1233687666+UOWHF_Add_c;
   		UOWHF_Add_c.3:=UOWHF_Result[3].31;
   		UOWHF_Result[3].31:=0;
   		UOWHF_Result[4]:=UOWHF_Result[4] + 279379632+UOWHF_Add_c;
   		UOWHF_Add_c.4:=UOWHF_Result[4].31;
   		UOWHF_Result[4].31:=0;
   		UOWHF_Result[5]:=UOWHF_Result[5] + 877536146+UOWHF_Add_c;
   		UOWHF_Add_c.5:=UOWHF_Result[5].31;
   		UOWHF_Result[5].31:=0;
   		UOWHF_Result[6]:=UOWHF_Result[6] + 10772756+UOWHF_Add_c;
   		UOWHF_Add_c.6:=UOWHF_Result[6].31;
   		UOWHF_Result[6].31:=0;
   	End_If;
   	If UOWHF_Msg[10].[15] Then
   		UOWHF_Result[0]:=UOWHF_Result[0] + 2133351485+UOWHF_Add_c;
   		UOWHF_Add_c.0:=UOWHF_Result[0].31;
   		UOWHF_Result[0].31:=0;
   		UOWHF_Result[1]:=UOWHF_Result[1] + 1410976862+UOWHF_Add_c;
   		UOWHF_Add_c.1:=UOWHF_Result[1].31;
   		UOWHF_Result[1].31:=0;
   		UOWHF_Result[2]:=UOWHF_Result[2] + 638097786+UOWHF_Add_c;
   		UOWHF_Add_c.2:=UOWHF_Result[2].31;
   		UOWHF_Result[2].31:=0;
   		UOWHF_Result[3]:=UOWHF_Result[3] + 1402702863+UOWHF_Add_c;
   		UOWHF_Add_c.3:=UOWHF_Result[3].31;
   		UOWHF_Result[3].31:=0;
   		UOWHF_Result[4]:=UOWHF_Result[4] + 563350383+UOWHF_Add_c;
   		UOWHF_Add_c.4:=UOWHF_Result[4].31;
   		UOWHF_Result[4].31:=0;
   		UOWHF_Result[5]:=UOWHF_Result[5] + 1243279963+UOWHF_Add_c;
   		UOWHF_Add_c.5:=UOWHF_Result[5].31;
   		UOWHF_Result[5].31:=0;
   		UOWHF_Result[6]:=UOWHF_Result[6] + 603841301+UOWHF_Add_c;
   		UOWHF_Add_c.6:=UOWHF_Result[6].31;
   		UOWHF_Result[6].31:=0;
   	End_If;
   	If UOWHF_Msg[10].[16] Then
   		UOWHF_Result[0]:=UOWHF_Result[0] + 1527964575+UOWHF_Add_c;
   		UOWHF_Add_c.0:=UOWHF_Result[0].31;
   		UOWHF_Result[0].31:=0;
   		UOWHF_Result[1]:=UOWHF_Result[1] + 1558705617+UOWHF_Add_c;
   		UOWHF_Add_c.1:=UOWHF_Result[1].31;
   		UOWHF_Result[1].31:=0;
   		UOWHF_Result[2]:=UOWHF_Result[2] + 204548494+UOWHF_Add_c;
   		UOWHF_Add_c.2:=UOWHF_Result[2].31;
   		UOWHF_Result[2].31:=0;
   		UOWHF_Result[3]:=UOWHF_Result[3] + 1124551983+UOWHF_Add_c;
   		UOWHF_Add_c.3:=UOWHF_Result[3].31;
   		UOWHF_Result[3].31:=0;
   		UOWHF_Result[4]:=UOWHF_Result[4] + 1720960624+UOWHF_Add_c;
   		UOWHF_Add_c.4:=UOWHF_Result[4].31;
   		UOWHF_Result[4].31:=0;
   		UOWHF_Result[5]:=UOWHF_Result[5] + 279739409+UOWHF_Add_c;
   		UOWHF_Add_c.5:=UOWHF_Result[5].31;
   		UOWHF_Result[5].31:=0;
   		UOWHF_Result[6]:=UOWHF_Result[6] + 946667469+UOWHF_Add_c;
   		UOWHF_Add_c.6:=UOWHF_Result[6].31;
   		UOWHF_Result[6].31:=0;
   	End_If;
   	If UOWHF_Msg[10].[17] Then
   		UOWHF_Result[0]:=UOWHF_Result[0] + 1919231123+UOWHF_Add_c;
   		UOWHF_Add_c.0:=UOWHF_Result[0].31;
   		UOWHF_Result[0].31:=0;
   		UOWHF_Result[1]:=UOWHF_Result[1] + 15594614+UOWHF_Add_c;
   		UOWHF_Add_c.1:=UOWHF_Result[1].31;
   		UOWHF_Result[1].31:=0;
   		UOWHF_Result[2]:=UOWHF_Result[2] + 999985952+UOWHF_Add_c;
   		UOWHF_Add_c.2:=UOWHF_Result[2].31;
   		UOWHF_Result[2].31:=0;
   		UOWHF_Result[3]:=UOWHF_Result[3] + 42612244+UOWHF_Add_c;
   		UOWHF_Add_c.3:=UOWHF_Result[3].31;
   		UOWHF_Result[3].31:=0;
   		UOWHF_Result[4]:=UOWHF_Result[4] + 733848970+UOWHF_Add_c;
   		UOWHF_Add_c.4:=UOWHF_Result[4].31;
   		UOWHF_Result[4].31:=0;
   		UOWHF_Result[5]:=UOWHF_Result[5] + 1382192730+UOWHF_Add_c;
   		UOWHF_Add_c.5:=UOWHF_Result[5].31;
   		UOWHF_Result[5].31:=0;
   		UOWHF_Result[6]:=UOWHF_Result[6] + 592381110+UOWHF_Add_c;
   		UOWHF_Add_c.6:=UOWHF_Result[6].31;
   		UOWHF_Result[6].31:=0;
   	End_If;
   	If UOWHF_Msg[10].[18] Then
   		UOWHF_Result[0]:=UOWHF_Result[0] + 722751617+UOWHF_Add_c;
   		UOWHF_Add_c.0:=UOWHF_Result[0].31;
   		UOWHF_Result[0].31:=0;
   		UOWHF_Result[1]:=UOWHF_Result[1] + 1707034784+UOWHF_Add_c;
   		UOWHF_Add_c.1:=UOWHF_Result[1].31;
   		UOWHF_Result[1].31:=0;
   		UOWHF_Result[2]:=UOWHF_Result[2] + 650598304+UOWHF_Add_c;
   		UOWHF_Add_c.2:=UOWHF_Result[2].31;
   		UOWHF_Result[2].31:=0;
   		UOWHF_Result[3]:=UOWHF_Result[3] + 980685617+UOWHF_Add_c;
   		UOWHF_Add_c.3:=UOWHF_Result[3].31;
   		UOWHF_Result[3].31:=0;
   		UOWHF_Result[4]:=UOWHF_Result[4] + 1531818986+UOWHF_Add_c;
   		UOWHF_Add_c.4:=UOWHF_Result[4].31;
   		UOWHF_Result[4].31:=0;
   		UOWHF_Result[5]:=UOWHF_Result[5] + 1899920054+UOWHF_Add_c;
   		UOWHF_Add_c.5:=UOWHF_Result[5].31;
   		UOWHF_Result[5].31:=0;
   		UOWHF_Result[6]:=UOWHF_Result[6] + 1081227376+UOWHF_Add_c;
   		UOWHF_Add_c.6:=UOWHF_Result[6].31;
   		UOWHF_Result[6].31:=0;
   	End_If;
   	If UOWHF_Msg[10].[19] Then
   		UOWHF_Result[0]:=UOWHF_Result[0] + 449851847+UOWHF_Add_c;
   		UOWHF_Add_c.0:=UOWHF_Result[0].31;
   		UOWHF_Result[0].31:=0;
   		UOWHF_Result[1]:=UOWHF_Result[1] + 1806679337+UOWHF_Add_c;
   		UOWHF_Add_c.1:=UOWHF_Result[1].31;
   		UOWHF_Result[1].31:=0;
   		UOWHF_Result[2]:=UOWHF_Result[2] + 1598159391+UOWHF_Add_c;
   		UOWHF_Add_c.2:=UOWHF_Result[2].31;
   		UOWHF_Result[2].31:=0;
   		UOWHF_Result[3]:=UOWHF_Result[3] + 2124828541+UOWHF_Add_c;
   		UOWHF_Add_c.3:=UOWHF_Result[3].31;
   		UOWHF_Result[3].31:=0;
   		UOWHF_Result[4]:=UOWHF_Result[4] + 804731841+UOWHF_Add_c;
   		UOWHF_Add_c.4:=UOWHF_Result[4].31;
   		UOWHF_Result[4].31:=0;
   		UOWHF_Result[5]:=UOWHF_Result[5] + 1250808565+UOWHF_Add_c;
   		UOWHF_Add_c.5:=UOWHF_Result[5].31;
   		UOWHF_Result[5].31:=0;
   		UOWHF_Result[6]:=UOWHF_Result[6] + 568554721+UOWHF_Add_c;
   		UOWHF_Add_c.6:=UOWHF_Result[6].31;
   		UOWHF_Result[6].31:=0;
   	End_If;
   	If UOWHF_Msg[10].[20] Then
   		UOWHF_Result[0]:=UOWHF_Result[0] + 247736158+UOWHF_Add_c;
   		UOWHF_Add_c.0:=UOWHF_Result[0].31;
   		UOWHF_Result[0].31:=0;
   		UOWHF_Result[1]:=UOWHF_Result[1] + 943808217+UOWHF_Add_c;
   		UOWHF_Add_c.1:=UOWHF_Result[1].31;
   		UOWHF_Result[1].31:=0;
   		UOWHF_Result[2]:=UOWHF_Result[2] + 120283341+UOWHF_Add_c;
   		UOWHF_Add_c.2:=UOWHF_Result[2].31;
   		UOWHF_Result[2].31:=0;
   		UOWHF_Result[3]:=UOWHF_Result[3] + 787622105+UOWHF_Add_c;
   		UOWHF_Add_c.3:=UOWHF_Result[3].31;
   		UOWHF_Result[3].31:=0;
   		UOWHF_Result[4]:=UOWHF_Result[4] + 1220909387+UOWHF_Add_c;
   		UOWHF_Add_c.4:=UOWHF_Result[4].31;
   		UOWHF_Result[4].31:=0;
   		UOWHF_Result[5]:=UOWHF_Result[5] + 1787946938+UOWHF_Add_c;
   		UOWHF_Add_c.5:=UOWHF_Result[5].31;
   		UOWHF_Result[5].31:=0;
   		UOWHF_Result[6]:=UOWHF_Result[6] + 2006270010+UOWHF_Add_c;
   		UOWHF_Add_c.6:=UOWHF_Result[6].31;
   		UOWHF_Result[6].31:=0;
   	End_If;
   	If UOWHF_Msg[10].[21] Then
   		UOWHF_Result[0]:=UOWHF_Result[0] + 1942854871+UOWHF_Add_c;
   		UOWHF_Add_c.0:=UOWHF_Result[0].31;
   		UOWHF_Result[0].31:=0;
   		UOWHF_Result[1]:=UOWHF_Result[1] + 2048257208+UOWHF_Add_c;
   		UOWHF_Add_c.1:=UOWHF_Result[1].31;
   		UOWHF_Result[1].31:=0;
   		UOWHF_Result[2]:=UOWHF_Result[2] + 944836520+UOWHF_Add_c;
   		UOWHF_Add_c.2:=UOWHF_Result[2].31;
   		UOWHF_Result[2].31:=0;
   		UOWHF_Result[3]:=UOWHF_Result[3] + 2026820467+UOWHF_Add_c;
   		UOWHF_Add_c.3:=UOWHF_Result[3].31;
   		UOWHF_Result[3].31:=0;
   		UOWHF_Result[4]:=UOWHF_Result[4] + 711914668+UOWHF_Add_c;
   		UOWHF_Add_c.4:=UOWHF_Result[4].31;
   		UOWHF_Result[4].31:=0;
   		UOWHF_Result[5]:=UOWHF_Result[5] + 1970053166+UOWHF_Add_c;
   		UOWHF_Add_c.5:=UOWHF_Result[5].31;
   		UOWHF_Result[5].31:=0;
   		UOWHF_Result[6]:=UOWHF_Result[6] + 1404598976+UOWHF_Add_c;
   		UOWHF_Add_c.6:=UOWHF_Result[6].31;
   		UOWHF_Result[6].31:=0;
   	End_If;
   	If UOWHF_Msg[10].[22] Then
   		UOWHF_Result[0]:=UOWHF_Result[0] + 907576588+UOWHF_Add_c;
   		UOWHF_Add_c.0:=UOWHF_Result[0].31;
   		UOWHF_Result[0].31:=0;
   		UOWHF_Result[1]:=UOWHF_Result[1] + 704377331+UOWHF_Add_c;
   		UOWHF_Add_c.1:=UOWHF_Result[1].31;
   		UOWHF_Result[1].31:=0;
   		UOWHF_Result[2]:=UOWHF_Result[2] + 526056233+UOWHF_Add_c;
   		UOWHF_Add_c.2:=UOWHF_Result[2].31;
   		UOWHF_Result[2].31:=0;
   		UOWHF_Result[3]:=UOWHF_Result[3] + 746855707+UOWHF_Add_c;
   		UOWHF_Add_c.3:=UOWHF_Result[3].31;
   		UOWHF_Result[3].31:=0;
   		UOWHF_Result[4]:=UOWHF_Result[4] + 1632965203+UOWHF_Add_c;
   		UOWHF_Add_c.4:=UOWHF_Result[4].31;
   		UOWHF_Result[4].31:=0;
   		UOWHF_Result[5]:=UOWHF_Result[5] + 1706158590+UOWHF_Add_c;
   		UOWHF_Add_c.5:=UOWHF_Result[5].31;
   		UOWHF_Result[5].31:=0;
   		UOWHF_Result[6]:=UOWHF_Result[6] + 367112835+UOWHF_Add_c;
   		UOWHF_Add_c.6:=UOWHF_Result[6].31;
   		UOWHF_Result[6].31:=0;
   	End_If;
   	If UOWHF_Msg[10].[23] Then
   		UOWHF_Result[0]:=UOWHF_Result[0] + 794882974+UOWHF_Add_c;
   		UOWHF_Add_c.0:=UOWHF_Result[0].31;
   		UOWHF_Result[0].31:=0;
   		UOWHF_Result[1]:=UOWHF_Result[1] + 1559202796+UOWHF_Add_c;
   		UOWHF_Add_c.1:=UOWHF_Result[1].31;
   		UOWHF_Result[1].31:=0;
   		UOWHF_Result[2]:=UOWHF_Result[2] + 533597257+UOWHF_Add_c;
   		UOWHF_Add_c.2:=UOWHF_Result[2].31;
   		UOWHF_Result[2].31:=0;
   		UOWHF_Result[3]:=UOWHF_Result[3] + 761339219+UOWHF_Add_c;
   		UOWHF_Add_c.3:=UOWHF_Result[3].31;
   		UOWHF_Result[3].31:=0;
   		UOWHF_Result[4]:=UOWHF_Result[4] + 1443683584+UOWHF_Add_c;
   		UOWHF_Add_c.4:=UOWHF_Result[4].31;
   		UOWHF_Result[4].31:=0;
   		UOWHF_Result[5]:=UOWHF_Result[5] + 498780807+UOWHF_Add_c;
   		UOWHF_Add_c.5:=UOWHF_Result[5].31;
   		UOWHF_Result[5].31:=0;
   		UOWHF_Result[6]:=UOWHF_Result[6] + 1184050969+UOWHF_Add_c;
   		UOWHF_Add_c.6:=UOWHF_Result[6].31;
   		UOWHF_Result[6].31:=0;
   	End_If;
   	If UOWHF_Msg[10].[24] Then
   		UOWHF_Result[0]:=UOWHF_Result[0] + 1715361051+UOWHF_Add_c;
   		UOWHF_Add_c.0:=UOWHF_Result[0].31;
   		UOWHF_Result[0].31:=0;
   		UOWHF_Result[1]:=UOWHF_Result[1] + 503936956+UOWHF_Add_c;
   		UOWHF_Add_c.1:=UOWHF_Result[1].31;
   		UOWHF_Result[1].31:=0;
   		UOWHF_Result[2]:=UOWHF_Result[2] + 934254333+UOWHF_Add_c;
   		UOWHF_Add_c.2:=UOWHF_Result[2].31;
   		UOWHF_Result[2].31:=0;
   		UOWHF_Result[3]:=UOWHF_Result[3] + 1253967563+UOWHF_Add_c;
   		UOWHF_Add_c.3:=UOWHF_Result[3].31;
   		UOWHF_Result[3].31:=0;
   		UOWHF_Result[4]:=UOWHF_Result[4] + 115833520+UOWHF_Add_c;
   		UOWHF_Add_c.4:=UOWHF_Result[4].31;
   		UOWHF_Result[4].31:=0;
   		UOWHF_Result[5]:=UOWHF_Result[5] + 1060993837+UOWHF_Add_c;
   		UOWHF_Add_c.5:=UOWHF_Result[5].31;
   		UOWHF_Result[5].31:=0;
   		UOWHF_Result[6]:=UOWHF_Result[6] + 1683624134+UOWHF_Add_c;
   		UOWHF_Add_c.6:=UOWHF_Result[6].31;
   		UOWHF_Result[6].31:=0;
   	End_If;
   	If UOWHF_Msg[10].[25] Then
   		UOWHF_Result[0]:=UOWHF_Result[0] + 1460646206+UOWHF_Add_c;
   		UOWHF_Add_c.0:=UOWHF_Result[0].31;
   		UOWHF_Result[0].31:=0;
   		UOWHF_Result[1]:=UOWHF_Result[1] + 895671635+UOWHF_Add_c;
   		UOWHF_Add_c.1:=UOWHF_Result[1].31;
   		UOWHF_Result[1].31:=0;
   		UOWHF_Result[2]:=UOWHF_Result[2] + 351368991+UOWHF_Add_c;
   		UOWHF_Add_c.2:=UOWHF_Result[2].31;
   		UOWHF_Result[2].31:=0;
   		UOWHF_Result[3]:=UOWHF_Result[3] + 1975753440+UOWHF_Add_c;
   		UOWHF_Add_c.3:=UOWHF_Result[3].31;
   		UOWHF_Result[3].31:=0;
   		UOWHF_Result[4]:=UOWHF_Result[4] + 1523645864+UOWHF_Add_c;
   		UOWHF_Add_c.4:=UOWHF_Result[4].31;
   		UOWHF_Result[4].31:=0;
   		UOWHF_Result[5]:=UOWHF_Result[5] + 1261931441+UOWHF_Add_c;
   		UOWHF_Add_c.5:=UOWHF_Result[5].31;
   		UOWHF_Result[5].31:=0;
   		UOWHF_Result[6]:=UOWHF_Result[6] + 1794091508+UOWHF_Add_c;
   		UOWHF_Add_c.6:=UOWHF_Result[6].31;
   		UOWHF_Result[6].31:=0;
   	End_If;
   	If UOWHF_Msg[10].[26] Then
   		UOWHF_Result[0]:=UOWHF_Result[0] + 618258893+UOWHF_Add_c;
   		UOWHF_Add_c.0:=UOWHF_Result[0].31;
   		UOWHF_Result[0].31:=0;
   		UOWHF_Result[1]:=UOWHF_Result[1] + 1637604100+UOWHF_Add_c;
   		UOWHF_Add_c.1:=UOWHF_Result[1].31;
   		UOWHF_Result[1].31:=0;
   		UOWHF_Result[2]:=UOWHF_Result[2] + 1304240362+UOWHF_Add_c;